(* Logix 5000 project; controller TemplateV1R0 vendor 1 type 14 code 222 rev 33.11; software revision 33.00; part 2 of 5 *)
(* tags used below, declared in another part *)
   EMs_Status : EquipmentModule[32];   // EquipmentModules information
   Sts_Clearing : BOOL;   // Clearing
   Sts_Aborting : BOOL;   // Aborting
   Sts_Aborted : BOOL;   // Aborted
   Sts_Resetting : BOOL;   // Resetting
   Sts_Production : BOOL;   // Machine is in production
   Sts_Maintenance : BOOL;   // Machine is in Maintenance
   Sts_Manual : BOOL;   // Machine is in Manual
   Sts_Cleaning : BOOL;   // Machine is in Cleaning
   Sts_MES : BOOL;   // Machine is in MES mode
   Sts_SemiAutomatic : BOOL;   // Machine is in Semi-Automatic
   PackTags : PACKMLv30;
   RecipeNumber : SINT;   // Recipe number selects which PackTag.command.product[#] will be used.
   DesignedSpeed : REAL;   // This tag represents the maximum design speed of the machine in primary packages per minute for the package configuration
   Sts_MachineFaulted : BOOL;   // Machine recieved an fault trigger
   MachineState : USINT;   // Technical Report Equipment States: 1 Clearing 2 Stopped 3 Starting 4 Idle 5 Suspended 6 Execute 7 Stopping 8 Aborting 9
   wrk_compare_UDINT : UDINT;
   cnf_EM_Size : DINT;   // size of array for equipmentmodules
   wrk_prev_state : DINT;   // local mem
   MachineMode : DINT;
   wrk_SwitchLayer_To_Cleaning : DINT;
   wrk_SwitchLayer_To_Maintenance : DINT;
   wrk_SwitchLayer_To_Manual : DINT;
   wrk_SwitchLayer_To_MES : DINT;
   wrk_SwitchLayer_To_Production : DINT;
   wrk_SwitchLayer_To_SemiAutomatic : DINT;
   T_second_puls : FBD_TIMER;   // local timer for just 1 second
   wrk_DateTime : LINT;
   T_ResetSignal_ON : FBD_TIMER;   // Local reset timer
   T_ResetSignal_HMI : FBD_TIMER;   // reset timer from HMI
   StateHistory : StateHistory[10];
(* ISA_TR_88_00_02, continued *)

   				15:	PackTags.Admin.StateCumulativeTime[MachineMode].Mode[15]	:=	PackTags.Admin.StateCumulativeTime[MachineMode].Mode[15]+1;
   				16:	PackTags.Admin.StateCumulativeTime[MachineMode].Mode[16]	:=	PackTags.Admin.StateCumulativeTime[MachineMode].Mode[16]+1;
   				17:	PackTags.Admin.StateCumulativeTime[MachineMode].Mode[17]	:=	PackTags.Admin.StateCumulativeTime[MachineMode].Mode[17]+1;
   				else
   				// undefined state.
   			end_case;
   		end_if;
   
   	#endregion
   
   	#region ProdConsumedCount
   		// should be done outsite of AOI, since the AOI cant keep track of this topic.
   	#endregion
   
   	#region ProdProcessedCount
   		// should be done outsite of AOI, since the AOI cant keep track of this topic.
   	#endregion
   
   	#region ProdDefectiveCount
   		// should be done outsite of AOI, since the AOI cant keep track of this topic.
   	#endregion
   
   	#region AccTimeSinceReset
   		if T_second_puls.DN then
   			if NOT Sts_Resetting then PackTags.Admin.AccTimeSinceReset:=PackTags.Admin.AccTimeSinceReset+1; end_if;		// count until machine has been in resetting.
   		end_if;
   		if T_ResetSignal_ON.TT OR T_ResetSignal_HMI.TT then PackTags.Admin.AccTimeSinceReset:=0; end_if;
   	#endregion
   
   	#region MachDesignSpeed
   		PackTags.Admin.MachDesignSpeed:=DesignedSpeed;
   	#endregion
   
   	#region PACDateTime
   	GSV(WallClockTime,,CurrentValue,wrk_DateTime);
   		#region PACDateTime.Date
   			PackTags.Admin.PACDateTime.Date:=wrk_DateTime;
   		#endregion
   		#region PACDateTime.Time
   			PackTags.Admin.PACDateTime.Time:=wrk_DateTime;
   		#endregion
   	#endregion
   #endregion
   #region HMI data representation
   	if StateHistory[0].State_Num <> MachineState then
   		for i := 1 to 9 do
   			StateHistory[10-i].State_Num 			:= StateHistory[9-i].State_Num;
   			StateHistory[10-i].Time_Spend_in_State 	:= StateHistory[9-i].Time_Spend_in_State;
   			StateHistory[10-i].Time_enteringState 	:= StateHistory[9-i].Time_enteringState;
   		end_for;
   		StateHistory[0].State_Num			:=MachineState;
   		StateHistory[0].Time_enteringState	:=wrk_DateTime;
   	end_if;
   	StateHistory[0].Time_Spend_in_State	:=PackTags.Admin.StateCurrentTime[MachineMode].Mode[MachineState];
   #endregion
END_ROUTINE

ROUTINE Prescan   (* structured text *)
// Clear old mem
   ////////////////////////////////////////////////////////////
   //   Copyright (c)
   //------------------------------------------------------------
   //   Routine: Prescan
   //   Author: WPI\tom.reit
   //   Created: 2-11-2022
   //------------------------------------------------------------
   //   Description:
   //           Clear old mem
   //
   //
   //   History:
   //
   ////////////////////////////////////////////////////////////
   #region EquipmentModule status
   	for i := 0 to 31 do
   		EMs_Status[i].Selected:=0;
   	end_for;
   #endregion
   wrk_compare_UDINT:=0;
   for i := 0 to 31 do
   	wrk_compare_UDINT:=(1*2**i)+wrk_compare_UDINT;	// set compare value, cant move 64bits so have to do some clever bit manipulation.
   end_for;
   SIZE(EMs_Status,0,cnf_EM_Size);
   cnf_EM_Size:=cnf_EM_Size-1;			// scale down because arrays start at 0
   
   
   wrk_prev_state						:=	-1;					// set mem state to something that machineState can never be. therfor the whileloop will always execute
   MachineState						:=	9;					// always start safe, in aborted.
   PackTags.Status.StateRequested		:=	MachineState;		// Set requested state same as actual state.
   
   wrk_SwitchLayer_To_Cleaning			:=0;		// Set layer switching to begin step.
   wrk_SwitchLayer_To_Maintenance		:=0;		// Set layer switching to begin step.
   wrk_SwitchLayer_To_Manual			:=0;		// Set layer switching to begin step.
   wrk_SwitchLayer_To_MES				:=0;		// Set layer switching to begin step.
   wrk_SwitchLayer_To_Production		:=0;		// Set layer switching to begin step.
   wrk_SwitchLayer_To_SemiAutomatic	:=0;		// Set layer switching to begin step.
   
   RecipeNumber						:=1;		// always run with first recipe on start.
   
   /* Reset ModeCumulativeTime for admin tags */
   for i := 0 to 6 do
   	PackTags.Admin.ModeCumulativeTime[i]:=0;
   end_for;
END_ROUTINE
END_ADD_ON_INSTRUCTION

ADD_ON_INSTRUCTION PF525_V3   (* revision 1.0 *)
// based on packml_V2_R1
VAR_INPUT
   PF_In : AB:PowerFlex525V_E_BBC69E8D:I:0;   // Powerflex object
   PF_Out : AB:PowerFlex525V_EENET_Drive:O:0;   // Powerflex object
END_VAR
VAR_IN_OUT
   Unit : ISA_TR_88_00_02; {required}   // Powerflex uses PackML for mode control
END_VAR
VAR_INPUT
   cnf_MinSpeed : REAL; {visible}   // Min speed the drive may run at
   cnf_MaxSpeed : REAL; {visible}   // Max speed the drive may run at
   cnf_MinHZ : REAL; {visible}   // max freq the drive may run at
   cnf_MaxHZ : REAL; {visible}   // max freq the drive may run at
   cnf_Direction : DINT; {visible}   // 0 = FWD 1 = REV
   Speed : REAL; {visible}   // required speed of drive. in units defined by user.
   Start : BOOL; {visible}   // Start the drive with Speed
END_VAR
VAR_OUTPUT
   Sts_Faulted : BOOL; {access Read Only, visible}   // Drive faulted, requires reset
   Sts_Drive_Running : BOOL; {access Read Only, visible}   // Motor is running
   Sts_Accelerating : BOOL; {access Read Only, visible}   // Drive is accelerating
   Sts_Execute : BOOL; {access Read Only, visible}   // motor is running at setpoint
   Sts_Decelerating : BOOL; {access Read Only, visible}   // Drive is decelerating
   Sts_Drive_Stopped : BOOL; {access Read Only, visible}   // Motor is NOT running
END_VAR
VAR_INPUT
   Reset : BOOL; {required}   // Reset drive signal resetting drive will only effect the AOI while drive is faulted
END_VAR
VAR_OUTPUT
   ActualSpeed : REAL; {access Read Only, visible}   // Feedback from drive what speed the drive is running at in user units
   Sts_DriveState : DINT; {access Read Only, visible}   // Drive states for HMI 0=Drive not active 1=Drive active 2=Spare 3=Manual turned on 4=Faulted
END_VAR
VAR_INPUT
   Force_On : BOOL; {visible}   // Turn drive on in manual & SemiAutomatic
   Force_Off : BOOL; {visible}   // Turn drive off in manual & SemiAutomatic
END_VAR
VAR_OUTPUT
   HMI_Show_Button : BOOL; {visible}
END_VAR
VAR
   ScaleSP : SCALE; {access None}   // scaling speed for drive
   TRUE : BOOL; {access None}   // macro to use TRUE
   FALSE : BOOL; {access None}   // Macro to use FALSE
   ons_Reset : FBD_ONESHOT; {access None}   // oneshot for resetting drive
   wrk_color : SINT; {access None}   // local mem for color of drive
   Build_Upper_Tag_AOI : Generate_HMI_Tag; {access None}
   Sts_Upper_Tag : STRING; {access Read Only}
   wrk_AddonName : STRING; {access None}
   GetLowerTag : Substring; {access None}
   Sts_Lower_Tag : STRING; {access Read Only}
   Sts_Show_HMIControls : BOOL;   // Show controls
END_VAR

ROUTINE Logic   (* structured text *)
// based on packml_V2_R1
   ////////////////////////////////////////////////////////////
   //   Copyright (c)
   //------------------------------------------------------------
   //   Routine: PF525_V3 - Logic
   //   Author: WPI\tom.reit
   //   Created: 17-11-2022
   //------------------------------------------------------------
   //   Description:
   //           based on packml_V2_R1
   //
   //
   //   History:
   //
   ////////////////////////////////////////////////////////////
   #region Macros
   	TRUE	:=1;																		// Mapped True macro
   	FALSE	:=0;																		// Mapped False macro
   	if cnf_Direction > 1 then cnf_Direction := 1; end_if;								// Prevent wrong direction input
   	if 0 > cnf_Direction then cnf_Direction := 0; end_if;								// Prevent wrong direction input
   #endregion
   #region Drive faulted & resetting it
   	if PF_In.Faulted AND NOT Reset then													// check if drive is faulted based on tags from PF525.
   		Sts_Faulted	:=	TRUE;															// Set drive faulted to true.
   		PF_Out.Stop	:= 	TRUE;															// Set Stop Drive to true.
   		PF_Out.Start:=	FALSE;															// Remove Start signal from drive.
   
   	elsif PF_In.Faulted AND Reset then													// check if drive is faulted based on tags from PF525 and reset signal is set.
   		PF_Out.ClearFaults	:=	TRUE;													// Set reset signal high for powerflex, this unlatches once the drive is back to its normal state.
   		Sts_Faulted			:=	FALSE;													// Set drive faulted to false.
   		PF_Out.Stop			:= 	FALSE;													// Set Stop Drive to false.
   	elsif PF_Out.ClearFaults AND NOT Reset then											// Check if PF_Out.ClearFaults is set.
   		if NOT PF_In.Faulted then														// Check if Drive is no longer faulted. waiting for drive to give feedback
   			PF_Out.ClearFaults	:= FALSE;												// Unlatch reset signal since reset was succesful.
   		end_if;
   	end_if;
   #endregion
   #region Start/Stop drive signal
   	if (Start AND NOT Force_Off) OR Force_On then															// Check if drive has start signal
   		#region Direction drive
   			if 	 cnf_Direction = 0 then 												// Check users input.
   					PF_Out.Reverse	:=	FALSE;											// Set direction of drive.
   					PF_Out.Forward	:=	TRUE;											// Set direction of drive.
   			elsif cnf_Direction = 1 then 												// Check users input.
   					PF_Out.Reverse	:=	TRUE;											// Set direction of drive.
   					PF_Out.Forward	:=	FALSE;											// Set direction of drive.
   			end_if;
   		#endregion
   		#region Start drive
   			if 	 	PF_Out.Stop		then PF_Out.Stop	:=FALSE; 	end_if;				// set stop drive to false.
   			if NOT	PF_Out.Start 	then PF_Out.Start	:=TRUE; 	end_if;				// Set Start drive to true.
   			#region Drive speed
   				ScaleSP.In			:=Speed;											// move speed to scale object.
   				PF_Out.FreqCommand	:=(ScaleSP.Out*100);								// convert to mili hz.
   			#endregion
   		#endregion
   	else																				// Check if drive has NO start signal
   		#region Stop drive
   			if 		PF_Out.Start 	then PF_Out.Start	:=FALSE; 	end_if;				// set Start drive to false.
   			if NOT 	PF_Out.Stop		then PF_Out.Stop	:=TRUE; 	end_if;				// set stop drive to True.
   			PF_Out.FreqCommand		:=0;												// Set speed of drive back to 0.
   		#endregion
   	end_if;
   #endregion
   #region Scale userinput
   	ScaleSP.In			:=Speed;														// Move speed into Scale object.
   	SCL(ScaleSP);																		// Scale Object.
   	ScaleSP.InEUMax		:=cnf_MaxHZ;													// Set Scale limits
   	ScaleSP.InEUMin		:=cnf_MinHZ;													// Set Scale limits
   	ScaleSP.InRawMax	:=cnf_MaxSpeed;													// Set Scale limits
   	ScaleSP.InRawMin	:=cnf_MinSpeed;													// Set Scale limits
   	ActualSpeed			:=(cnf_MaxSpeed/cnf_MaxHZ) * (PF_In.OutputFreq/100);			// Convert powerflex feedback frequenty to user units.
   #endregion
   
   #region Feedback to user about drive.
   	if PF_In.Accelerating 	then 	Sts_Accelerating	:=	TRUE; 	else 	Sts_Accelerating	:=	FALSE; 	end_if;
   	if PF_In.Decelerating 	then	Sts_Decelerating	:=	TRUE;	else	Sts_Decelerating	:=	FALSE;	end_if;
   	if PF_In.Faulted		then	Sts_Faulted			:=	TRUE;	else	Sts_Faulted			:=	FALSE;	end_if;
   	if PF_In.Active			then	Sts_Drive_Running	:=	TRUE;	else	Sts_Drive_Running	:=	FALSE;	end_if;
   	if PF_In.OutputFreq<>0	then	Sts_Drive_Stopped	:=	FALSE; 											end_if;
   	if PF_In.OutputFreq =0	then	Sts_Drive_Stopped	:=	TRUE; 											end_if;
   	if PF_In.AtReference	then	Sts_Execute			:=	TRUE;	else	Sts_Execute			:=	FALSE;	end_if;
   	#region HMI Drive color.
   	/*
   		Colortable:
   		0:drive is not active	(grey)
   		1:drive is active		(green)
   		2:forced on				(blue)
   		3:forced off			(white)
   	*/
   		#region Select drive state
   			if Sts_Drive_Stopped 					   			then Sts_DriveState:=0; end_if;
   			if Sts_Drive_Running AND (Start	AND NOT Force_On)	then Sts_DriveState:=1; end_if;
   			if Sts_Drive_Running AND Force_On					then Sts_DriveState:=2; end_if;
   			if (Start AND Force_Off AND Unit.Sts_SemiAutomatic)	then Sts_DriveState:=3; end_if;
   		#endregion
   	#endregion
   #endregion
   
   if s:fs then
   	Generate_HMI_Tag(Build_Upper_Tag_AOI,Sts_Upper_Tag);
   	GSV(Routine,THIS,Name,wrk_AddonName);
   	Substring(GetLowerTag,wrk_AddonName,7,wrk_AddonName.LEN,Sts_Lower_Tag);
   end_if;
   
   if NOT (Unit.Sts_SemiAutomatic OR Unit.Sts_Manual) then
   	Force_Off:=FALSE;
   	Force_On:=FALSE;
   end_if;
   
   if Unit.Sts_SemiAutomatic OR Unit.Sts_Manual then
   	HMI_Show_Button:=TRUE;
   Else
   	HMI_Show_Button:=FALSE;
   end_if;
END_ROUTINE
END_ADD_ON_INSTRUCTION

ADD_ON_INSTRUCTION Phase_Call   (* revision 1.0, ExecuteEnableInFalse *)
VAR_IN_OUT
   Phase : PhaseObject; {required}
END_VAR
VAR_OUTPUT
   PhaseCall_Enabled : BOOL; {access Read Only, visible}   // Phase is enabled
   PhaseCall_Faulted : BOOL; {access Read Only, visible}   // Phase is faulted
   PhaseCall_Ownership : BOOL; {access Read Only, visible}   // Phase is executing
   EN : BOOL; {access Read Only, visible}   // Phase is enabled
   IP : BOOL; {access Read Only, visible}   // Phase is in proces / Active
   ER : BOOL; {access Read Only, visible}   // Phase is faulted
   PC : BOOL; {access Read Only, visible}   // Phase is completed
   FLAGS : INT; {access Read Only, visible}   // Status
        .1   // PhaseCall_Enabled
        .2   // PhaseCall_Faulted
        .3   // PhaseCall_Ownership
        .4   // PhaseHandler_Enabled
        .5   // PhaseHandler_InProces
        .6   // PhaseHandler_ProcesComplete
        .7   // PhaseHandler_Execute
END_VAR
VAR_INPUT
   Reset : BOOL; {visible}   // Reset PhaseCall outputs & Flags
   cnf_DisableAutomaticReset : BOOL := 1;   // Resets PC & ER automaticly if phasecall is not enabled
END_VAR
VAR
   Wrk_Call_Name : STRING[3] := ([0] := 'Procedure_Batter', [1] := 'Unit1_Procedural_Model', [2] := 'CIP'); {access None}
   wrk_TotalName : STRING; {access None}
   i : INT; {access None}   // index num
   wrk_Insert_Start_Pos : DINT; {access None}   // local var
   Sts_TotalName : STRING := 'Procedure_Batter -> Unit1_Procedural_Model -> UP_CIP_PH_FillingColdWater'; {access None}   // total name of phasecall Task -> Program -> Routine
   SEQ_TakeOwnership : DINT; {access None}   // Take ownership of a phase.
   wrk_tempName : STRING; {access None}
   wrk_Flags : DINT; {access None}   // local flags memory
END_VAR

ROUTINE EnableInFalse   (* structured text *)
   ////////////////////////////////////////////////////////////
   //   Copyright (c)
   //------------------------------------------------------------
   //   Routine: EnableInFalse
   //   Author: WPI\tom.reit
   //   Created: 1-2-2023
   //------------------------------------------------------------
   //   Description:
   //
   //
   //   History:
   //
   ////////////////////////////////////////////////////////////
   #region Reset phasecall outputs & Flags
   	if Reset OR (wrk_Flags<>FLAGS) then
   		FLAGS		:=0;
   		EN			:=0;
   		IP			:=0;
   		ER			:=0;
   		PC			:=0;
   		wrk_Flags	:=FLAGS;
   		Reset		:=0;
   	end_if;
   #endregion
   if Phase.PhaseHandler.Sts_Locked AND PhaseCall_Ownership then
   	PhaseCall_Enabled	:=0;
   	PhaseCall_Ownership	:=1;			// holding ownership signal while phasehandler is releasing lock.
   	Phase.PhaseHandler.Req_Unlock:=1;	// set unlock signal, phasehandler will unlock.
   	SEQ_TakeOwnership:=4;				// Pre-set fault if same instruction gets scanned twice move to error state.
   	#region Copy phase status to local outputs
   		EN:=Phase.Status.EN;
   		IP:=Phase.Status.IP;
   		ER:=Phase.Status.ER;
   		PC:=Phase.Status.PC;
   	#endregion
   else
   	PhaseCall_Enabled	:=0;			//
   	SEQ_TakeOwnership	:=0;			//
   	PhaseCall_Ownership	:=0;			//
   	#region Copy phase status to local outputs
   		EN:=0;
   		IP:=0;
   		if cnf_DisableAutomaticReset then
   			/* Currently disabled, since we want to keep track of the last states. */
   			// ER:=0;
   			// PC:=0;
   		else
   			ER:=0;
   			PC:=0;
   		end_if;
   	#endregion
   end_if;
   
   
END_ROUTINE

ROUTINE Logic   (* structured text *)
   ////////////////////////////////////////////////////////////
   //   Copyright (c)
   //------------------------------------------------------------
   //   Routine: PhaseCall - Logic
   //   Author: WPI\tom.reit
   //   Created: 1-2-2023
   //------------------------------------------------------------
   //   Description:
   //
   //
   //   History:
   //
   ////////////////////////////////////////////////////////////
   #region Reset phasecall outputs & Flags
   	if Reset then
   		FLAGS	:=0;
   		EN		:=0;
   		IP		:=0;
   		ER		:=0;
   		PC		:=0;
   		Reset	:=0;
   	end_if;
   #endregion
   
   if EnableIn then
   	PhaseCall_Enabled:=1;
   	case SEQ_TakeOwnership of
   		0: // Step 0, Send request to Phase_Handler.
   			Phase.PhaseHandler.Req_Lock		:=1;												// Set lock reques to phase_handler
   			SEQ_TakeOwnership				:=1;												// Move to next state.
   		1: // Step 1, wait for handshake from Phase_Handler.
   			if NOT Phase.PhaseHandler.Req_Lock 			then SEQ_TakeOwnership:=2; end_if;		// wait for feedback
   		2: // Step 2, Acknowledge.
   			Sts_TotalName:='|';														// clear previous data
   			GSV(Program,THIS,Name,Wrk_Call_Name[0]);								// Get program name
   			GSV(Routine,THIS,Name,Wrk_Call_Name[1]);								// Get Routine name
   
   			#region owner string
   				wrk_Insert_Start_Pos:=Wrk_Call_Name[0].LEN+1;
   				INSERT(Wrk_Call_Name[0],Sts_TotalName,wrk_Insert_Start_Pos,Wrk_Call_Name[0]);
   				INSERT(Wrk_Call_Name[1],Wrk_Call_Name[0],1,wrk_tempName);
   				INSERT(wrk_tempName,Sts_TotalName,1,Sts_TotalName);
   			#endregion
   			if Phase.PhaseHandler.Sts_Accept_lock 		then SEQ_TakeOwnership:=3; end_if;		// Phase was succesfully assigned
   			if NOT Phase.PhaseHandler.Sts_Accept_lock 	then SEQ_TakeOwnership:=4; end_if;		// Phase was already locked, go to an error state.
   		3: // Succesfull lock
   			Phase.Status.Owner:=Sts_TotalName;
   			PhaseCall_Ownership:=1;																	// in ownership
   			PhaseCall_Faulted:=0;																	// No errors
   
   			#region Copy phase status to local outputs
   				EN:=Phase.Status.EN;
   				IP:=Phase.Status.IP;
   				ER:=Phase.Status.ER;
   				PC:=Phase.Status.PC;
   			#endregion
   
   
   			if NOT Phase.PhaseHandler.Sts_Locked  		then SEQ_TakeOwnership:=4;	end_if;		// if for some reason the phase gets unlocked go to error state since phase has not been succesfully executed.
   		4: // Faulted
   			PhaseCall_Faulted:=1;																	// No errors		// Error
   		else
   			SEQ_TakeOwnership:=0;
   	end_case;
   end_if;
   
   #region Flags
   	FLAGS.0:=PhaseCall_Enabled;
   	FLAGS.1:=PhaseCall_Faulted;
   	FLAGS.2:=PhaseCall_Ownership;
   	FLAGS.3:=EN;
   	FLAGS.4:=IP;
   	FLAGS.5:=ER;
   	FLAGS.6:=PC;
   	FLAGS.7:=Phase.PhaseHandler.Sts_Execute;
   	wrk_Flags:=FLAGS;
   #endregion
END_ROUTINE
END_ADD_ON_INSTRUCTION

ADD_ON_INSTRUCTION Phase_Handler   (* revision 1.0, ExecutePrescan *)
VAR_IN_OUT
   Phase_Status : PhaseStatus; {required}
END_VAR
VAR_OUTPUT
   Sts_Locked : BOOL; {access Read Only, visible}   // Phase is executing and locked
END_VAR
VAR_INPUT
   Req_Lock : BOOL;   // Operation locks phase
END_VAR
VAR_OUTPUT
   Sts_Accept_lock : BOOL; {access Read Only}   // Lock signal is accepted by handler
END_VAR
VAR_INPUT
   Req_Unlock : BOOL;   // if Phase is locked, only owner can send unlock.
END_VAR
VAR_OUTPUT
   Sts_Execute : BOOL; {access Read Only, visible}   // Phase may execute
END_VAR
VAR_INPUT
   Force_Unlock : BOOL; {visible}   // Forces an unlock and phase may be reassigned. keep in mind the phasecall that was in process will move to an error state.
END_VAR
VAR_OUTPUT
   Sts_AssignTime : LINT; {access Read Only, visible}
   Sts_UnassignTime : LINT; {access Read Only, visible}
END_VAR
VAR_INPUT
   Watchdog : BOOL;
END_VAR
VAR_OUTPUT
   Sts_Unlocking : BOOL; {access Read Only, visible}   // Phase recieved an unlock request and is waiting for IP to go LOW.
END_VAR
VAR
   wrk_lockState : BOOL; {access None}   // local mem
   wrk_Instance : DINT; {access None}
   lock_ID : LINT; {access None}   // based on when lock was succesfull
END_VAR

ROUTINE Logic   (* structured text *)
   ////////////////////////////////////////////////////////////
   //   Copyright (c)
   //------------------------------------------------------------
   //   Routine: Phase_Handler - Logic
   //   Author: WPI\tom.reit
   //   Created: 1-2-2023
   //------------------------------------------------------------
   //   Description:
   //
   //
   //   History:
   //
   ////////////////////////////////////////////////////////////
   #region Prevent user from unlatching/latching Lock Status
   	wrk_lockState:=Sts_Locked;
   	Sts_Locked:=wrk_lockState;
   #endregion
   #region Request lock and assign phase
   	if Req_Lock AND NOT Sts_Locked then
   		GSV(WallClockTime,,CurrentValue,Sts_AssignTime);
   		GSV(Routine,THIS,INSTANCE,wrk_Instance);
   		GSV(WallClockTime,,CurrentValue,lock_ID);
   		Sts_UnassignTime:=0;	// remove unasign time
   		Req_Lock		:=0;	// handshake to Phase_call
   		Sts_Accept_lock	:=1;	// accept lock
   		Sts_Locked		:=1;	// accept lock
   		Sts_Execute		:=1;	// Set phase to execute
   	end_if;
   #endregion
   #region Deal with request lock while phase was allready assigned.
   	if Req_Lock AND Sts_Locked then
   		Req_Lock		:=0;	// handshake to Phase_call
   		Sts_Accept_lock	:=0;	// decline lock
   	end_if;
   
   #endregion
   #region Force unlock
   	if Force_Unlock then
   		Req_Unlock		:=1;
   		Force_Unlock	:=0;
   	end_if;
   #endregion
   #region Unassign phase and unlock phase
   	if Req_Unlock AND Sts_Locked then
   		Sts_Execute:=0;
   		Sts_Unlocking:=1;
   		if NOT Phase_Status.IP then
   			GSV(WallClockTime,,CurrentValue,Sts_UnassignTime);
   			Sts_Locked:=0;
   			Sts_Unlocking:=0;
   			Req_Unlock:=0;
   		end_if;
   	end_if;
   #endregion
   #region Set phase to execute/running
   	if Sts_Locked then
   		Phase_Status.EN:=1;
   	else
   		Phase_Status.EN:=0;
   	end_if;
   #endregion
   
   if NOT Sts_Execute then Phase_Status.CurrentAction:=''; end_if;
END_ROUTINE

ROUTINE Prescan   (* structured text *)
   ////////////////////////////////////////////////////////////
   //   Copyright (c)
   //------------------------------------------------------------
   //   Routine: Prescan
   //   Author: WPI\tom.reit
   //   Created: 2-2-2023
   //------------------------------------------------------------
   //   Description:
   //
   //
   //   History:
   //
   ////////////////////////////////////////////////////////////
   Watchdog			:=0;
   Sts_Accept_lock		:=0;
   Sts_AssignTime		:=0;
   Sts_Locked			:=0;
   Sts_Execute			:=0;
   Sts_UnassignTime	:=0;
END_ROUTINE
END_ADD_ON_INSTRUCTION

ADD_ON_INSTRUCTION PID_V3   (* revision 1.0, ExecutePrescan *)
// using an Infinite impulse response filter for the derivative
VAR_INPUT
   Enable_PID : BOOL; {visible}   // Turn on the PID controller
   cnf_setPID_Values : BOOL; {visible}
   cnf_Use_PID : SINT := 7; {visible}   // P is always acitve bit 0 = P bit 1 = I bit 2 = D
   Kp : REAL; {visible}   // Proportional
   Ki : REAL; {visible}   // Integral
   Kd : REAL; {visible}   // Derivative
   N : REAL; {visible}   // Filter constant
   dt : REAL; {visible}   // update time
   setpoint : REAL; {visible}
   measured_value : REAL; {visible}
END_VAR
VAR_OUTPUT
   actuator_value : REAL; {access Read Only, visible}   // current actuator value
END_VAR
VAR_INPUT
   HandValue : REAL; {visible}   // Static handvalue
END_VAR
VAR_OUTPUT
   Output : REAL; {access Read Only, visible}
   tau : REAL; {access Read Only}
   alpha : REAL; {access Read Only}
END_VAR
VAR
   A0 : REAL; {access None}
   A1 : REAL; {access None}
   error : REAL[3]; {access None}
   A0d : REAL; {access None}
   A1d : REAL; {access None}
   A2d : REAL; {access None}
   fd1 : REAL; {access None}
   fd0 : REAL; {access None}
   d1 : REAL; {access None}
   d0 : REAL; {access None}
   time_interval : FBD_TIMER; {access None}
   proportional : REAL; {access None}
   wrk_output : REAL; {access Read Only}
   wrk_kp : REAL; {access None}   // local mem
   wrk_ki : REAL; {access None}   // local mem
   wrk_kd : REAL; {access None}   // local mem
   wrk_dt : REAL; {access None}   // local mem
   wrk_N : REAL; {access None}   // local mem
END_VAR

ROUTINE Logic   (* structured text *)
// using an Infinite impulse response filter for the derivative
   ////////////////////////////////////////////////////////////
   //   Copyright (c)
   //------------------------------------------------------------
   //   Routine: PID_V3 - Logic
   //   Author: WPI\tom.reit
   //   Created: 2-12-2022
   //------------------------------------------------------------
   //   Description:
   //           using an Infinite impulse response filter for the
   //           derivative
   //
   //
   //   History:
   //
   ////////////////////////////////////////////////////////////
   #region Timer (dt)
   	time_interval.TimerEnable:=Enable_PID;
   	TONR(time_interval);
   	time_interval.Reset:=0;
   	time_interval.PRE:=dt*1000;
   #endregion
   #region Startup PID
   if Kp <> wrk_kp then cnf_setPID_Values:=1; wrk_kp:=Kp; end_if;
   if Ki <> wrk_ki then cnf_setPID_Values:=1; wrk_ki:=Ki; end_if;
   if Kd <> wrk_kd then cnf_setPID_Values:=1; wrk_kd:=Kd; end_if;
   if dt <> wrk_dt then cnf_setPID_Values:=1; wrk_dt:=dt; end_if;
   if N  <> wrk_N  then cnf_setPID_Values:=1; wrk_N :=N;  end_if;
   
   	if cnf_setPID_Values AND Enable_PID then
   		A0 := Kp + Ki*dt;
   		A1 := 0-Kp;
   		error[2] := 0; // e(t-2)
   		error[1] := 0; // e(t-1)
   		error[0] := 0; // e(t)
   		Output := actuator_value;  // Usually the current value of the actuator
   		A0d:= Kd/dt;
   		A1d:= (0- 2.0)*Kd/dt;
   		A2d:= Kd/dt;
   		N := N;
   		tau := Kd / (Kp*N); // IIR filter time constant
   		alpha:= dt / (2*tau);
   		d0 := 0;
   		d1 := 0;
   		fd0 := 0;
   		fd1 := 0;
   		if NOT cnf_Use_PID.0 then cnf_Use_PID.0 := 1; end_if;// makesure P is always active.
   		cnf_setPID_Values:=0;
   	end_if;
   
   #endregion
   #region PID logic, constant loop
   	if time_interval.DN then
   	    error[2] := error[1];
   	    error[1] := error[0];
   	    error[0] := setpoint - measured_value;
   		wrk_output:=Output;
   
   		case cnf_Use_PID of
   			0: cnf_Use_PID:=1;
   			1: // P 	controller
   				proportional := error[0];
   				wrk_output := Kp * proportional;
   			3: // PI 	controller
   				wrk_output := wrk_output + A0 * error[0] + A1 * error[1];
   			5: // PD 	controller
   				proportional := error[0];
   				wrk_output := Kp * proportional;
   				d1 := d0;
   			    d0 := A0d * error[0] + A1d * error[1] + A2d * error[2];
   			    fd1 := fd0;
   			    fd0 := ((alpha) / (alpha + 1)) * (d0 + d1) - ((alpha - 1) / (alpha + 1)) * fd1;
   			    wrk_output := wrk_output + fd0;
   			7: // PID 	controller
   				wrk_output := wrk_output + A0 * error[0] + A1 * error[1];
   			    d1 := d0;
   			    d0 := A0d * error[0] + A1d * error[1] + A2d * error[2];
   			    fd1 := fd0;
   			    fd0 := ((alpha) / (alpha + 1)) * (d0 + d1) - ((alpha - 1) / (alpha + 1)) * fd1;
   			    wrk_output := wrk_output + fd0;
   			else
   				cnf_Use_PID:=1;
   		end_case;
   		if wrk_output>=100 then wrk_output:=100; end_if;
   		if 0>=wrk_output then wrk_output:=0; end_if;
   		Output:=wrk_output;
   		time_interval.Reset:=1;
   	end_if;
   #endregion
   #region PID Handvalue
   	if NOT Enable_PID then
   		Output:=HandValue;
   	end_if;
   #endregion
END_ROUTINE

ROUTINE Prescan   (* structured text *)
   ////////////////////////////////////////////////////////////
   //   Copyright (c)
   //------------------------------------------------------------
   //   Routine: Prescan
   //   Author: WPI\tom.reit
   //   Created: 5-12-2022
   //------------------------------------------------------------
   //   Description:
   //
   //
   //   History:
   //
   ////////////////////////////////////////////////////////////
   wrk_dt :=0;
   wrk_kd :=0;
   wrk_ki :=0;
   wrk_kp :=0;
   wrk_N  :=0;
   wrk_output :=0;
END_ROUTINE
END_ADD_ON_INSTRUCTION

ADD_ON_INSTRUCTION PILZ_GuardSwitch   (* revision 1.0, ExecutePrescan *)
// based on model 21904-3FR-03 PSEN sl-0.5p
VAR_INPUT
   I_DoorClosed : BOOL := 1; {required}   // Y32 door is closed
END_VAR
VAR_OUTPUT
   O_LockDoor : BOOL; {required}   // signal to lock door S31
END_VAR
VAR_INPUT
   I_Doorlocked_S1 : BOOL; {required}   // 12
   I_Doorlocked_S2 : BOOL; {required}   // 22
END_VAR
VAR_OUTPUT
   DoorLocked : BOOL := 1; {visible}   // door is locked and feedback signals are OK
   Faulted : BOOL; {visible}   // Something went verie vrong much problem many oplossingen zoeken
   DoorClosed : BOOL; {visible}   // Door is closed
   DoorOpen : BOOL; {visible}   // Door is open
END_VAR
VAR_INPUT
   HMI_Request_LockDoor : BOOL; {visible}   // user requests to lock the door
   Reset : BOOL; {required}   // reset pilz logic
   OEM_Force_Open : BOOL := 1; {visible}   // Simulates tank door locked & Closed
END_VAR
VAR
   T_DetectDoorClosed : TIMER := (PRE := 500); {access None}
   T_wrk_LockingTime : TIMER := (PRE := 500); {access None}
   cnf_Hold_lock_In_Fault : BOOL := 1; {access None}   // config, hold lock when faulted. only lets go of lock once reset has been pressed.
END_VAR

ROUTINE Logic   (* ladder *)
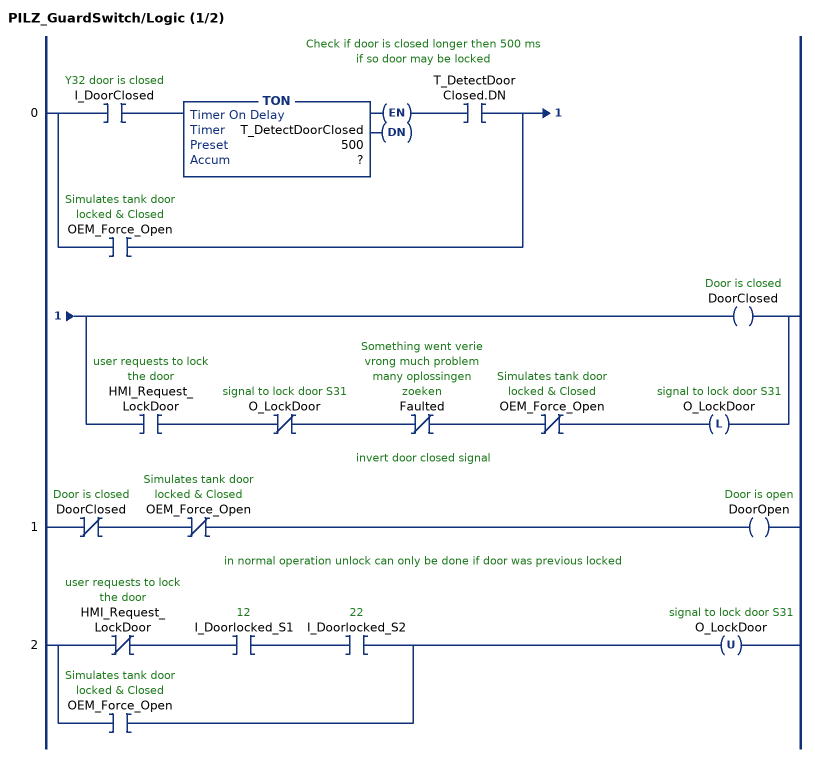
   // Check if door is closed longer then 500 ms
   // if so door may be locked
   0: [XIC(I_DoorClosed) TON(T_DetectDoorClosed,?,?) XIC(T_DetectDoorClosed.DN) ,XIC(OEM_Force_Open) ][OTE(DoorClosed) ,XIC(HMI_Request_LockDoor) XIO(O_LockDoor) XIO(Faulted) XIO(OEM_Force_Open) OTL(O_LockDoor) ];
   // invert door closed signal
   1: XIO(DoorClosed)XIO(OEM_Force_Open)OTE(DoorOpen);
   // in normal operation unlock can only be done if door was previous locked
   2: [XIO(HMI_Request_LockDoor) XIC(I_Doorlocked_S1) XIC(I_Doorlocked_S2) ,XIC(OEM_Force_Open) ]OTU(O_LockDoor);
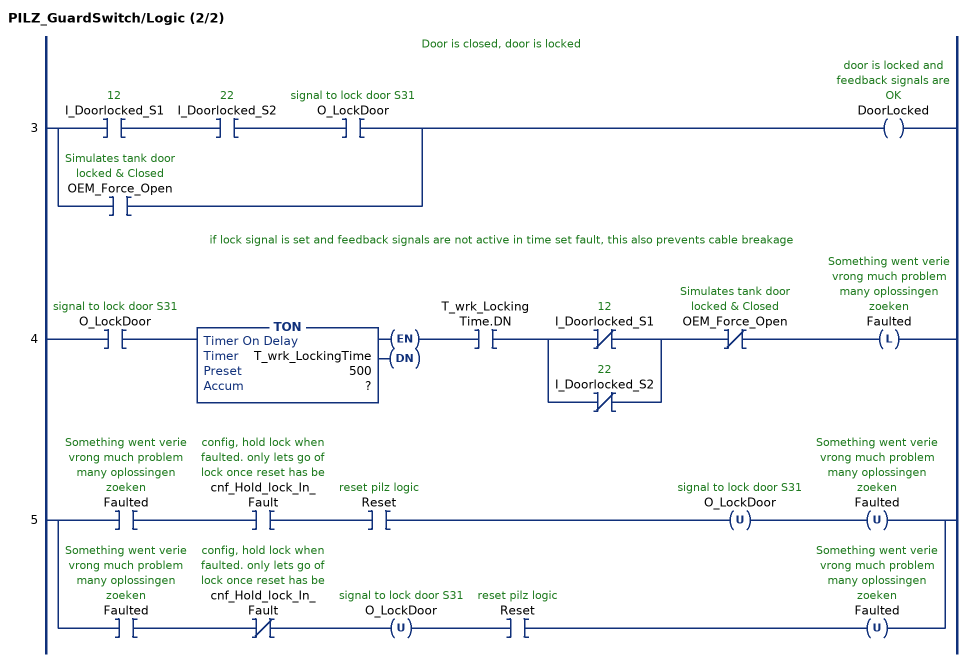
   // Door is closed, door is locked
   3: [XIC(I_Doorlocked_S1) XIC(I_Doorlocked_S2) XIC(O_LockDoor) ,XIC(OEM_Force_Open) ]OTE(DoorLocked);
   // if lock signal is set and feedback signals are not active in time set fault, this also prevents cable breakage
   4: XIC(O_LockDoor)TON(T_wrk_LockingTime,?,?)XIC(T_wrk_LockingTime.DN)[XIO(I_Doorlocked_S1) ,XIO(I_Doorlocked_S2) ]XIO(OEM_Force_Open)OTL(Faulted);
   5: [XIC(Faulted) XIC(cnf_Hold_lock_In_Fault) XIC(Reset) OTU(O_LockDoor) OTU(Faulted) ,XIC(Faulted) XIO(cnf_Hold_lock_In_Fault) OTU(O_LockDoor) XIC(Reset) OTU(Faulted) ];
END_ROUTINE

ROUTINE Prescan   (* structured text *)
   T_DetectDoorClosed.PRE	:=	500;
   T_wrk_LockingTime.PRE	:=	1000;
   cnf_Hold_lock_In_Fault 	:= 	0;
   OEM_Force_Open			:= 	0;
END_ROUTINE
END_ADD_ON_INSTRUCTION

ADD_ON_INSTRUCTION ServoMotor   (* revision 1.0, ExecutePrescan *)
VAR_IN_OUT
   Axis : AXIS_CIP_DRIVE; {required}
   Unit : ISA_TR_88_00_02; {required}
END_VAR
VAR_INPUT
   In_Enable : BOOL; {visible}   // Enable drive
   In_Disable : BOOL; {visible}
   In_Reset : BOOL; {visible}
   In_Home : BOOL; {visible}   // Home axis
   Force_ON : BOOL; {visible}   // Forces drive to enable
   Force_Off : BOOL; {visible}   // Forces drive to disable
END_VAR
VAR_OUTPUT
   Sts_DriveState : DINT;
   Sts_Faulted : BOOL; {visible}   // Drive faulted
   Sts_MotionError : BOOL; {visible}   // Motion instruciton faulted
   Sts_Enabled : BOOL := 1; {visible}   // Axis is enabled
   Sts_Disabled : BOOL; {visible}   // Axis is disabled
   Sts_Homing : BOOL; {visible}   // Axis is currently homing
   Sts_Homed : BOOL; {visible}   // Axis is homed
   HMI_Show_Button : BOOL;
END_VAR
VAR
   ons_ClearFlags : BOOL[32];   // local ons
   MC_MSO : MOTION_INSTRUCTION;
   MC_MSF : MOTION_INSTRUCTION; {access None}
   MC_MAFR : MOTION_INSTRUCTION; {access None}
   MC_MAH : MOTION_INSTRUCTION; {access None}
   Build_Upper_Tag_AOI : Generate_HMI_Tag; {access None}
   Sts_Upper_Tag : STRING;
   wrk_AddonName : STRING;
   Sts_Lower_Tag : STRING;
   GetLowerTag : Substring; {access None}
END_VAR

ROUTINE Logic   (* ladder *)
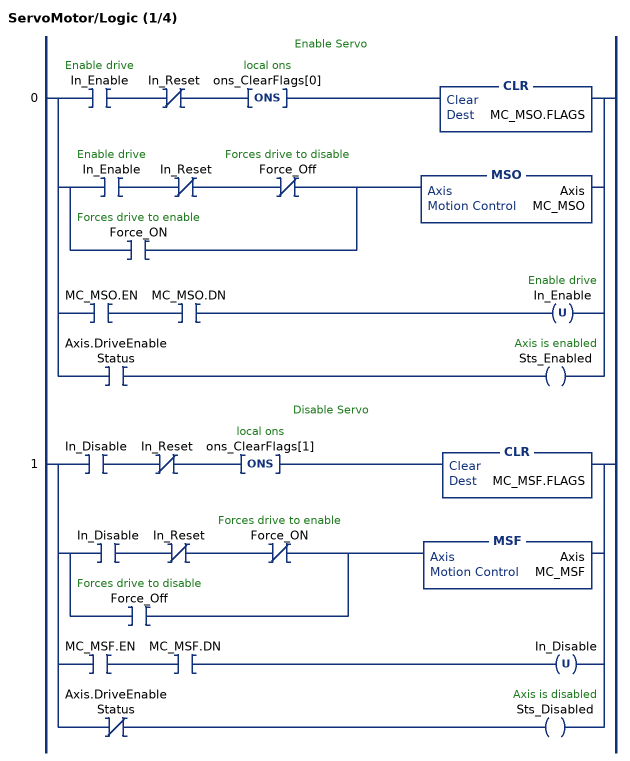
   // Enable Servo
   0: [XIC(In_Enable) XIO(In_Reset) ONS(ons_ClearFlags[0]) CLR(MC_MSO.FLAGS) ,[XIC(In_Enable) XIO(In_Reset) XIO(Force_Off) ,XIC(Force_ON) ] MSO(Axis,MC_MSO) ,XIC(MC_MSO.EN) XIC(MC_MSO.DN) OTU(In_Enable) ,XIC(Axis.DriveEnableStatus) OTE(Sts_Enabled) ];
   // Disable Servo
   1: [XIC(In_Disable) XIO(In_Reset) ONS(ons_ClearFlags[1]) CLR(MC_MSF.FLAGS) ,[XIC(In_Disable) XIO(In_Reset) XIO(Force_ON) ,XIC(Force_Off) ] MSF(Axis,MC_MSF) ,XIC(MC_MSF.EN) XIC(MC_MSF.DN) OTU(In_Disable) ,XIO(Axis.DriveEnableStatus) OTE(Sts_Disabled) ];
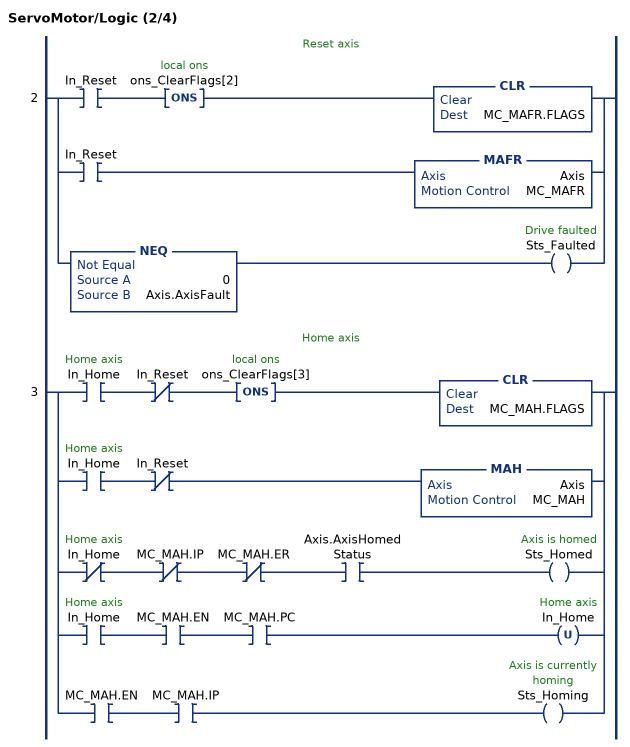
   // Reset axis
   2: [XIC(In_Reset) ONS(ons_ClearFlags[2]) CLR(MC_MAFR.FLAGS) ,XIC(In_Reset) MAFR(Axis,MC_MAFR) ,NEQ(0,Axis.AxisFault) OTE(Sts_Faulted) ];
   // Home axis
   3: [XIC(In_Home) XIO(In_Reset) ONS(ons_ClearFlags[3]) CLR(MC_MAH.FLAGS) ,XIC(In_Home) XIO(In_Reset) MAH(Axis,MC_MAH) ,XIO(In_Home) XIO(MC_MAH.IP) XIO(MC_MAH.ER) XIC(Axis.AxisHomedStatus) OTE(Sts_Homed) ,XIC(In_Home) XIC(MC_MAH.EN) XIC(MC_MAH.PC) OTU(In_Home) ,XIC(MC_MAH.EN) XIC(MC_MAH.IP) OTE(Sts_Homing) ];